// TIA Portal project "Sistema_de_silos" (V16) (continued)
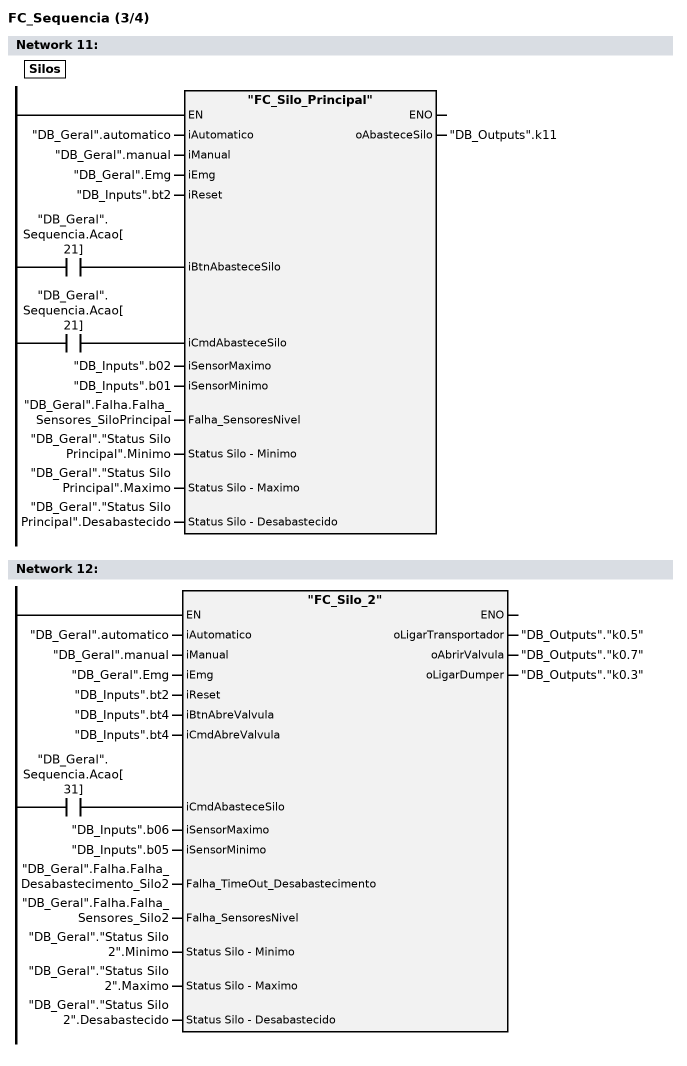
   Label( Silos )
   RUNG wire#powerrail
      "FC_Silo_Principal"(iBtnAbasteceSilo := wire#w1, iCmdAbasteceSilo := wire#w2, iAutomatico := "DB_Geral".automatico, iManual := "DB_Geral".manual, iEmg := "DB_Geral".Emg, iReset := "DB_Inputs".bt2, iSensorMaximo := "DB_Inputs".b02, iSensorMinimo := "DB_Inputs".b01, Falha_SensoresNivel := "DB_Geral".Falha.Falha_Sensores_SiloPrincipal, "Status Silo - Minimo" := "DB_Geral"."Status Silo Principal".Minimo, "Status Silo - Maximo" := "DB_Geral"."Status Silo Principal".Maximo, "Status Silo - Desabastecido" := "DB_Geral"."Status Silo Principal".Desabastecido, oAbasteceSilo => "DB_Outputs".k11)
   END_RUNG
   RUNG wire#powerrail
      Contact( "DB_Geral".Sequencia.Acao[21] )
   END_RUNG wire#w1
   RUNG wire#powerrail
      Contact( "DB_Geral".Sequencia.Acao[21] )
   END_RUNG wire#w2
   // the same network as SCL:
   Silos:
   "FC_Silo_Principal"(iAutomatico := "DB_Geral".automatico,
                       iManual := "DB_Geral".manual,
                       iEmg := "DB_Geral".Emg,
                       iReset := "DB_Inputs".bt2,
                       iBtnAbasteceSilo := "DB_Geral".Sequencia.Acao[21],
                       iCmdAbasteceSilo := "DB_Geral".Sequencia.Acao[21],
                       iSensorMaximo := "DB_Inputs".b02,
                       iSensorMinimo := "DB_Inputs".b01,
                       Falha_SensoresNivel := "DB_Geral".Falha.Falha_Sensores_SiloPrincipal,
                       "Status Silo - Minimo" := "DB_Geral"."Status Silo Principal".Minimo,
                       "Status Silo - Maximo" := "DB_Geral"."Status Silo Principal".Maximo,
                       "Status Silo - Desabastecido" := "DB_Geral"."Status Silo Principal".Desabastecido,
                       oAbasteceSilo => "DB_Outputs".k11);
END_REGION

REGION Network 12
   RUNG wire#powerrail
      "FC_Silo_2"(iCmdAbasteceSilo := wire#w1, iAutomatico := "DB_Geral".automatico, iManual := "DB_Geral".manual, iEmg := "DB_Geral".Emg, iReset := "DB_Inputs".bt2, iBtnAbreValvula := "DB_Inputs".bt4, iCmdAbreValvula := "DB_Inputs".bt4, iSensorMaximo := "DB_Inputs".b06, iSensorMinimo := "DB_Inputs".b05, Falha_TimeOut_Desabastecimento := "DB_Geral".Falha.Falha_Desabastecimento_Silo2, Falha_SensoresNivel := "DB_Geral".Falha.Falha_Sensores_Silo2, "Status Silo - Minimo" := "DB_Geral"."Status Silo 2".Minimo, "Status Silo - Maximo" := "DB_Geral"."Status Silo 2".Maximo, "Status Silo - Desabastecido" := "DB_Geral"."Status Silo 2".Desabastecido, oLigarTransportador => "DB_Outputs"."k0.5", oAbrirValvula => "DB_Outputs"."k0.7", oLigarDumper => "DB_Outputs"."k0.3")
   END_RUNG
   RUNG wire#powerrail
      Contact( "DB_Geral".Sequencia.Acao[31] )
   END_RUNG wire#w1
   // the same network as SCL:
   "FC_Silo_2"(iAutomatico := "DB_Geral".automatico,
               iManual := "DB_Geral".manual,
               iEmg := "DB_Geral".Emg,
               iReset := "DB_Inputs".bt2,
               iBtnAbreValvula := "DB_Inputs".bt4,
               iCmdAbreValvula := "DB_Inputs".bt4,
               iCmdAbasteceSilo := "DB_Geral".Sequencia.Acao[31],
               iSensorMaximo := "DB_Inputs".b06,
               iSensorMinimo := "DB_Inputs".b05,
               Falha_TimeOut_Desabastecimento := "DB_Geral".Falha.Falha_Desabastecimento_Silo2,
               Falha_SensoresNivel := "DB_Geral".Falha.Falha_Sensores_Silo2,
               "Status Silo - Minimo" := "DB_Geral"."Status Silo 2".Minimo,
               "Status Silo - Maximo" := "DB_Geral"."Status Silo 2".Maximo,
               "Status Silo - Desabastecido" := "DB_Geral"."Status Silo 2".Desabastecido,
               oLigarTransportador => "DB_Outputs"."k0.5",
               oAbrirValvula => "DB_Outputs"."k0.7",
               oLigarDumper => "DB_Outputs"."k0.3");
END_REGION

REGION Network 13
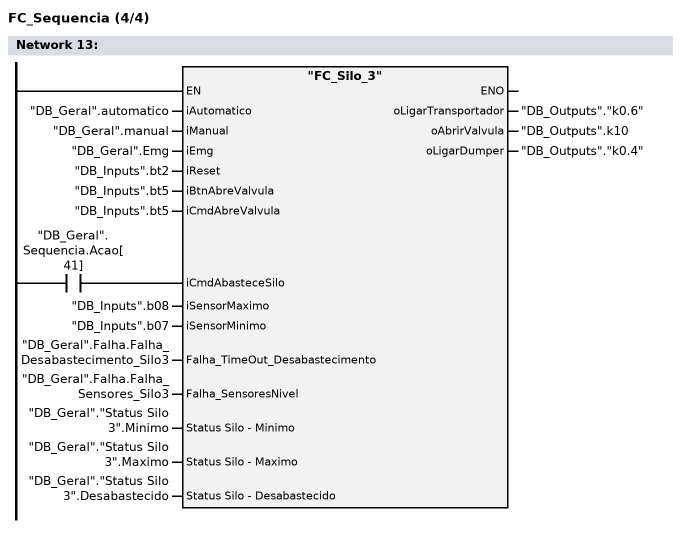
   RUNG wire#powerrail
      "FC_Silo_3"(iCmdAbasteceSilo := wire#w1, iAutomatico := "DB_Geral".automatico, iManual := "DB_Geral".manual, iEmg := "DB_Geral".Emg, iReset := "DB_Inputs".bt2, iBtnAbreValvula := "DB_Inputs".bt5, iCmdAbreValvula := "DB_Inputs".bt5, iSensorMaximo := "DB_Inputs".b08, iSensorMinimo := "DB_Inputs".b07, Falha_TimeOut_Desabastecimento := "DB_Geral".Falha.Falha_Desabastecimento_Silo3, Falha_SensoresNivel := "DB_Geral".Falha.Falha_Sensores_Silo3, "Status Silo - Minimo" := "DB_Geral"."Status Silo 3".Minimo, "Status Silo - Maximo" := "DB_Geral"."Status Silo 3".Maximo, "Status Silo - Desabastecido" := "DB_Geral"."Status Silo 3".Desabastecido, oLigarTransportador => "DB_Outputs"."k0.6", oAbrirValvula => "DB_Outputs".k10, oLigarDumper => "DB_Outputs"."k0.4")
   END_RUNG
   RUNG wire#powerrail
      Contact( "DB_Geral".Sequencia.Acao[41] )
   END_RUNG wire#w1
   // the same network as SCL:
   "FC_Silo_3"(iAutomatico := "DB_Geral".automatico,
               iManual := "DB_Geral".manual,
               iEmg := "DB_Geral".Emg,
               iReset := "DB_Inputs".bt2,
               iBtnAbreValvula := "DB_Inputs".bt5,
               iCmdAbreValvula := "DB_Inputs".bt5,
               iCmdAbasteceSilo := "DB_Geral".Sequencia.Acao[41],
               iSensorMaximo := "DB_Inputs".b08,
               iSensorMinimo := "DB_Inputs".b07,
               Falha_TimeOut_Desabastecimento := "DB_Geral".Falha.Falha_Desabastecimento_Silo3,
               Falha_SensoresNivel := "DB_Geral".Falha.Falha_Sensores_Silo3,
               "Status Silo - Minimo" := "DB_Geral"."Status Silo 3".Minimo,
               "Status Silo - Maximo" := "DB_Geral"."Status Silo 3".Maximo,
               "Status Silo - Desabastecido" := "DB_Geral"."Status Silo 3".Desabastecido,
               oLigarTransportador => "DB_Outputs"."k0.6",
               oAbrirValvula => "DB_Outputs".k10,
               oLigarDumper => "DB_Outputs"."k0.4");
END_REGION
END_FUNCTION

FUNCTION "FC_Silo_2" : Void   // FC5, LAD
{ S7_Optimized_Access := 'TRUE' }
VERSION : 0.1
   VAR_INPUT
      iAutomatico : Bool;
      iManual : Bool;
      iEmg : Bool;
      iReset : Bool;
      iBtnAbreValvula : Bool;
      iCmdAbreValvula : Bool;
      iCmdAbasteceSilo : Bool;
      iSensorMaximo : Bool;
      iSensorMinimo : Bool;
   END_VAR
   VAR_OUTPUT
      oLigarTransportador : Bool;
      oAbrirValvula : Bool;
      oLigarDumper : Bool;
   END_VAR
   VAR_IN_OUT
      Falha_TimeOut_Desabastecimento : Bool;
      Falha_SensoresNivel : Bool;
      "Status Silo - Minimo" : Bool;
      "Status Silo - Maximo" : Bool;
      "Status Silo - Desabastecido" : Bool;
   END_VAR
   VAR CONSTANT
      Velocidade_fluxo : Int := 12;
   END_VAR
BEGIN

REGION Network 1
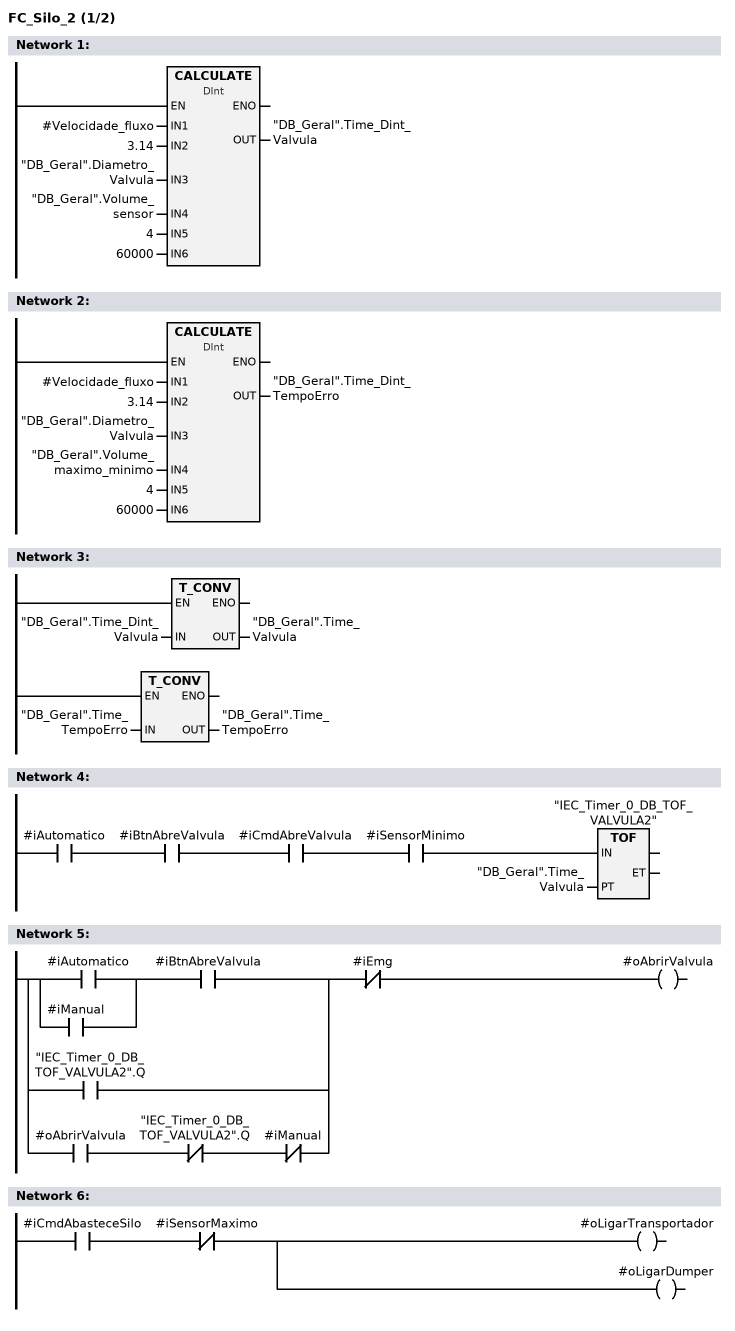
   RUNG wire#powerrail
      { S7_Templates := "SrcType := DInt"; S7_Expression := "(IN4 / (IN1* ((IN2*IN3*IN3) / IN5))) * IN6" } Calculate(in1 := #Velocidade_fluxo, in2 := 3.14, in3 := "DB_Geral".Diametro_Valvula, in4 := "DB_Geral".Volume_sensor, in5 := 4, in6 := 60000, out => "DB_Geral".Time_Dint_Valvula)
   END_RUNG
   // the same network as SCL:
   "DB_Geral".Time_Dint_Valvula := ("DB_Geral".Volume_sensor / (#Velocidade_fluxo* ((3.14*"DB_Geral".Diametro_Valvula*"DB_Geral".Diametro_Valvula) / 4))) * 60000;
END_REGION

REGION Network 2
   RUNG wire#powerrail
      { S7_Templates := "SrcType := DInt"; S7_Expression := "(IN4 / (IN1* ((IN2*IN3*IN3) / IN5))) * IN6" } Calculate(in1 := #Velocidade_fluxo, in2 := 3.14, in3 := "DB_Geral".Diametro_Valvula, in4 := "DB_Geral".Volume_maximo_minimo, in5 := 4, in6 := 60000, out => "DB_Geral".Time_Dint_TempoErro)
   END_RUNG
   // the same network as SCL:
   "DB_Geral".Time_Dint_TempoErro := ("DB_Geral".Volume_maximo_minimo / (#Velocidade_fluxo* ((3.14*"DB_Geral".Diametro_Valvula*"DB_Geral".Diametro_Valvula) / 4))) * 60000;
END_REGION

REGION Network 3
   "DB_Geral".Time_Valvula := T_CONV(IN := "DB_Geral".Time_Dint_Valvula);
   "DB_Geral".Time_TempoErro := T_CONV(IN := "DB_Geral".Time_TempoErro);
END_REGION

REGION Network 4
   "IEC_Timer_0_DB_TOF_VALVULA2".TOF(IN := #iAutomatico AND #iBtnAbreValvula AND #iCmdAbreValvula AND #iSensorMinimo,
                           PT := "DB_Geral".Time_Valvula);
END_REGION

REGION Network 5
   RUNG wire#powerrail
      Contact( #iAutomatico )
      wire#w1
      Contact( #iBtnAbreValvula )
      wire#w2
      I_Contact( #iEmg )
      Coil( #oAbrirValvula )
   END_RUNG
   RUNG wire#powerrail
      Contact( #iManual )
   END_RUNG wire#w1
   RUNG wire#powerrail
      Contact( "IEC_Timer_0_DB_TOF_VALVULA2".Q )
   END_RUNG wire#w2
   RUNG wire#powerrail
      Contact( #oAbrirValvula )
      I_Contact( "IEC_Timer_0_DB_TOF_VALVULA2".Q )
      I_Contact( #iManual )
   END_RUNG wire#w2
   // the same network as SCL:
   #oAbrirValvula := (((#iAutomatico OR #iManual) AND #iBtnAbreValvula) OR "IEC_Timer_0_DB_TOF_VALVULA2".Q OR (#oAbrirValvula AND NOT "IEC_Timer_0_DB_TOF_VALVULA2".Q AND NOT #iManual)) AND NOT #iEmg;
END_REGION

REGION Network 6
   RUNG wire#powerrail
      Contact( #iCmdAbasteceSilo )
      I_Contact( #iSensorMaximo )
      wire#w1
      Coil( #oLigarTransportador )
   END_RUNG
   RUNG wire#w1
      Coil( #oLigarDumper )
   END_RUNG
   // the same network as SCL:
   #oLigarTransportador := #iCmdAbasteceSilo AND NOT #iSensorMaximo;
   #oLigarDumper := #oLigarTransportador;
END_REGION

REGION Network 7: Silo Principal - Reserva do produto
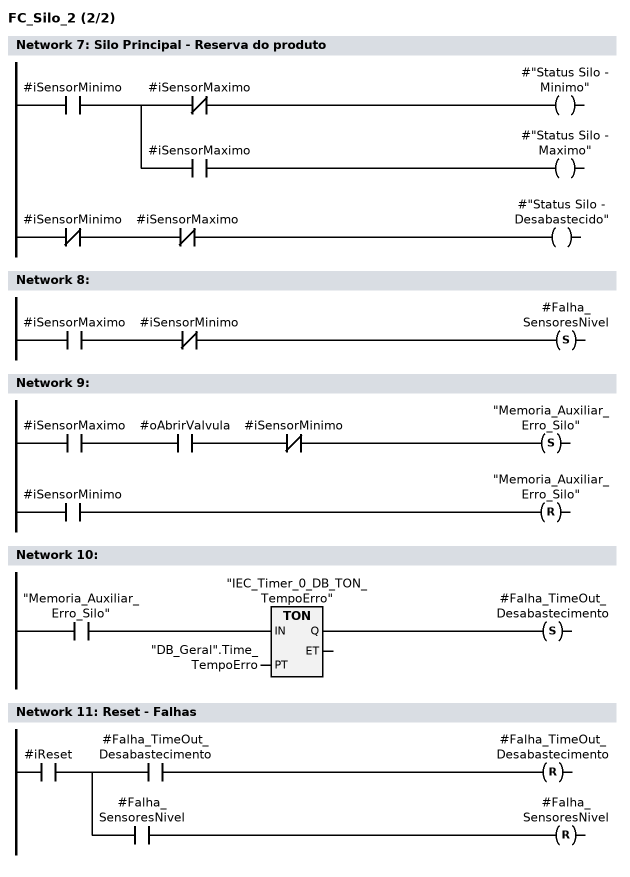
   RUNG wire#powerrail
      Contact( #iSensorMinimo )
      wire#w1
      I_Contact( #iSensorMaximo )
      Coil( #"Status Silo - Minimo" )
   END_RUNG
   RUNG wire#w1
      Contact( #iSensorMaximo )
      Coil( #"Status Silo - Maximo" )
   END_RUNG
   RUNG wire#powerrail
      I_Contact( #iSensorMinimo )
      I_Contact( #iSensorMaximo )
      Coil( #"Status Silo - Desabastecido" )
   END_RUNG
   // the same network as SCL:
   #"Status Silo - Minimo" := #iSensorMinimo AND NOT #iSensorMaximo;
   #"Status Silo - Maximo" := #iSensorMinimo AND #iSensorMaximo;
   #"Status Silo - Desabastecido" := NOT #iSensorMinimo AND NOT #iSensorMaximo;
END_REGION

REGION Network 8
   RUNG wire#powerrail
      Contact( #iSensorMaximo )
      I_Contact( #iSensorMinimo )
      S_Coil( #Falha_SensoresNivel )
   END_RUNG
   // the same network as SCL:
   IF #iSensorMaximo AND NOT #iSensorMinimo THEN #Falha_SensoresNivel := TRUE; END_IF;
END_REGION

REGION Network 9
   RUNG wire#powerrail
      Contact( #iSensorMaximo )
      Contact( #oAbrirValvula )
      I_Contact( #iSensorMinimo )
      S_Coil( "Memoria_Auxiliar_Erro_Silo" )
   END_RUNG
   RUNG wire#powerrail
      Contact( #iSensorMinimo )
      R_Coil( "Memoria_Auxiliar_Erro_Silo" )
   END_RUNG
   // the same network as SCL:
   IF #iSensorMaximo AND #oAbrirValvula AND NOT #iSensorMinimo THEN
       "Memoria_Auxiliar_Erro_Silo" := TRUE;
   END_IF;
   IF #iSensorMinimo THEN "Memoria_Auxiliar_Erro_Silo" := FALSE; END_IF;
END_REGION

REGION Network 10
   "IEC_Timer_0_DB_TON_TempoErro".TON(IN := "Memoria_Auxiliar_Erro_Silo", PT := "DB_Geral".Time_TempoErro);
   IF "IEC_Timer_0_DB_TON_TempoErro".Q THEN #Falha_TimeOut_Desabastecimento := TRUE; END_IF;
END_REGION

REGION Network 11: Reset - Falhas
   RUNG wire#powerrail
      Contact( #iReset )
      wire#w1
      Contact( #Falha_TimeOut_Desabastecimento )
      R_Coil( #Falha_TimeOut_Desabastecimento )
   END_RUNG
   RUNG wire#w1
      Contact( #Falha_SensoresNivel )
      R_Coil( #Falha_SensoresNivel )
   END_RUNG
   // the same network as SCL:
   IF #iReset AND #Falha_TimeOut_Desabastecimento THEN #Falha_TimeOut_Desabastecimento := FALSE; END_IF;
   IF #iReset AND #Falha_SensoresNivel THEN #Falha_SensoresNivel := FALSE; END_IF;
END_REGION
END_FUNCTION

FUNCTION "FC_Silo_Principal" : Void   // FC6, LAD
{ S7_Optimized_Access := 'TRUE' }
VERSION : 0.1
   VAR_INPUT
      iAutomatico : Bool;
      iManual : Bool;
      iEmg : Bool;
      iReset : Bool;
      iBtnAbasteceSilo : Bool;
      iCmdAbasteceSilo : Bool;
      iSensorMaximo : Bool;
      iSensorMinimo : Bool;
   END_VAR
   VAR_OUTPUT
      oAbasteceSilo : Bool;
   END_VAR
   VAR_IN_OUT
      Falha_SensoresNivel : Bool;
      "Status Silo - Minimo" : Bool;
      "Status Silo - Maximo" : Bool;
      "Status Silo - Desabastecido" : Bool;
   END_VAR
BEGIN

REGION Network 1
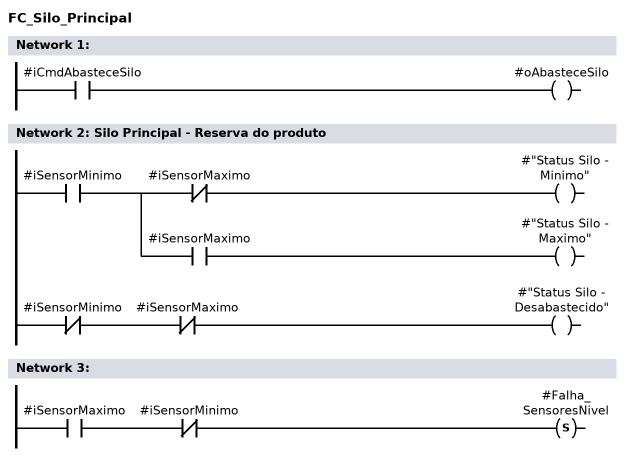
   RUNG wire#powerrail
      Contact( #iCmdAbasteceSilo )
      Coil( #oAbasteceSilo )
   END_RUNG
   // the same network as SCL:
   #oAbasteceSilo := #iCmdAbasteceSilo;
END_REGION

REGION Network 2: Silo Principal - Reserva do produto
   RUNG wire#powerrail
      Contact( #iSensorMinimo )
      wire#w1
      I_Contact( #iSensorMaximo )
      Coil( #"Status Silo - Minimo" )
   END_RUNG
   RUNG wire#w1
      Contact( #iSensorMaximo )
      Coil( #"Status Silo - Maximo" )
   END_RUNG
   RUNG wire#powerrail
      I_Contact( #iSensorMinimo )
      I_Contact( #iSensorMaximo )
      Coil( #"Status Silo - Desabastecido" )
   END_RUNG
   // the same network as SCL:
   #"Status Silo - Minimo" := #iSensorMinimo AND NOT #iSensorMaximo;
   #"Status Silo - Maximo" := #iSensorMinimo AND #iSensorMaximo;
   #"Status Silo - Desabastecido" := NOT #iSensorMinimo AND NOT #iSensorMaximo;
END_REGION

REGION Network 3
   RUNG wire#powerrail
      Contact( #iSensorMaximo )
      I_Contact( #iSensorMinimo )
      S_Coil( #Falha_SensoresNivel )
   END_RUNG
   // the same network as SCL:
   IF #iSensorMaximo AND NOT #iSensorMinimo THEN #Falha_SensoresNivel := TRUE; END_IF;
END_REGION
END_FUNCTION

FUNCTION "FC_Silo_3" : Void   // FC7, LAD
{ S7_Optimized_Access := 'TRUE' }
VERSION : 0.1
   VAR_INPUT
      iAutomatico : Bool;
      iManual : Bool;
      iEmg : Bool;
      iReset : Bool;
      iBtnAbreValvula : Bool;
      iCmdAbreValvula : Bool;
      iCmdAbasteceSilo : Bool;
      iSensorMaximo : Bool;
      iSensorMinimo : Bool;
   END_VAR
   VAR_OUTPUT
      oLigarTransportador : Bool;
      oAbrirValvula : Bool;
      oLigarDumper : Bool;
   END_VAR
   VAR_IN_OUT
      Falha_TimeOut_Desabastecimento : Bool;
      Falha_SensoresNivel : Bool;
      "Status Silo - Minimo" : Bool;
      "Status Silo - Maximo" : Bool;
      "Status Silo - Desabastecido" : Bool;
   END_VAR
   VAR CONSTANT
      Velocidade_fluxo : Int := 12;
   END_VAR
BEGIN

REGION Network 1
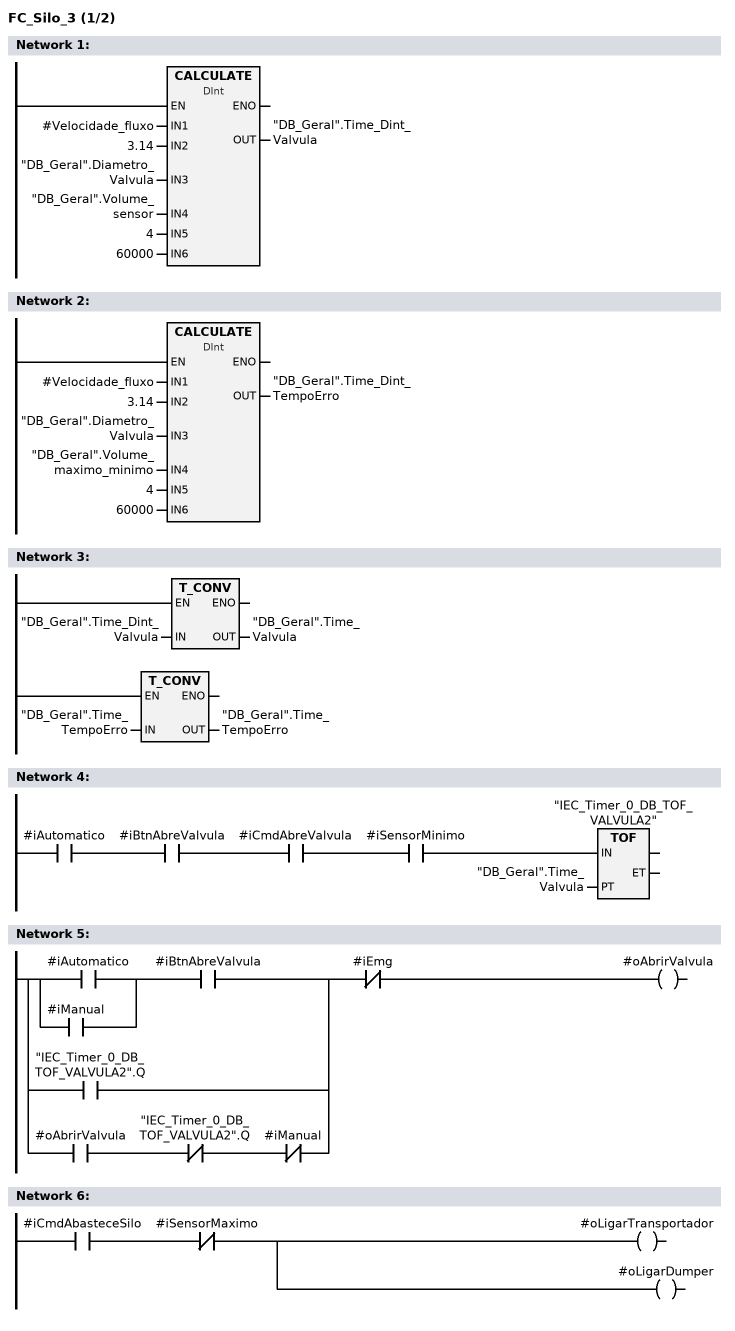
   RUNG wire#powerrail
      { S7_Templates := "SrcType := DInt"; S7_Expression := "(IN4 / (IN1* ((IN2*IN3*IN3) / IN5))) * IN6" } Calculate(in1 := #Velocidade_fluxo, in2 := 3.14, in3 := "DB_Geral".Diametro_Valvula, in4 := "DB_Geral".Volume_sensor, in5 := 4, in6 := 60000, out => "DB_Geral".Time_Dint_Valvula)
   END_RUNG
   // the same network as SCL:
   "DB_Geral".Time_Dint_Valvula := ("DB_Geral".Volume_sensor / (#Velocidade_fluxo* ((3.14*"DB_Geral".Diametro_Valvula*"DB_Geral".Diametro_Valvula) / 4))) * 60000;
END_REGION

REGION Network 2
   RUNG wire#powerrail
      { S7_Templates := "SrcType := DInt"; S7_Expression := "(IN4 / (IN1* ((IN2*IN3*IN3) / IN5))) * IN6" } Calculate(in1 := #Velocidade_fluxo, in2 := 3.14, in3 := "DB_Geral".Diametro_Valvula, in4 := "DB_Geral".Volume_maximo_minimo, in5 := 4, in6 := 60000, out => "DB_Geral".Time_Dint_TempoErro)
   END_RUNG
   // the same network as SCL:
   "DB_Geral".Time_Dint_TempoErro := ("DB_Geral".Volume_maximo_minimo / (#Velocidade_fluxo* ((3.14*"DB_Geral".Diametro_Valvula*"DB_Geral".Diametro_Valvula) / 4))) * 60000;
END_REGION

REGION Network 3
   "DB_Geral".Time_Valvula := T_CONV(IN := "DB_Geral".Time_Dint_Valvula);
   "DB_Geral".Time_TempoErro := T_CONV(IN := "DB_Geral".Time_TempoErro);
END_REGION

REGION Network 4
   "IEC_Timer_0_DB_TOF_VALVULA2".TOF(IN := #iAutomatico AND #iBtnAbreValvula AND #iCmdAbreValvula AND #iSensorMinimo,
                           PT := "DB_Geral".Time_Valvula);
END_REGION

REGION Network 5
   RUNG wire#powerrail
      Contact( #iAutomatico )
      wire#w1
      Contact( #iBtnAbreValvula )
      wire#w2
      I_Contact( #iEmg )
      Coil( #oAbrirValvula )
   END_RUNG
   RUNG wire#powerrail
      Contact( #iManual )
   END_RUNG wire#w1
   RUNG wire#powerrail
      Contact( "IEC_Timer_0_DB_TOF_VALVULA2".Q )
   END_RUNG wire#w2
   RUNG wire#powerrail
      Contact( #oAbrirValvula )
      I_Contact( "IEC_Timer_0_DB_TOF_VALVULA2".Q )
      I_Contact( #iManual )
   END_RUNG wire#w2
   // the same network as SCL:
   #oAbrirValvula := (((#iAutomatico OR #iManual) AND #iBtnAbreValvula) OR "IEC_Timer_0_DB_TOF_VALVULA2".Q OR (#oAbrirValvula AND NOT "IEC_Timer_0_DB_TOF_VALVULA2".Q AND NOT #iManual)) AND NOT #iEmg;
END_REGION

REGION Network 6
   RUNG wire#powerrail
      Contact( #iCmdAbasteceSilo )
      I_Contact( #iSensorMaximo )
      wire#w1
      Coil( #oLigarTransportador )
   END_RUNG
   RUNG wire#w1
      Coil( #oLigarDumper )
   END_RUNG
   // the same network as SCL:
   #oLigarTransportador := #iCmdAbasteceSilo AND NOT #iSensorMaximo;
   #oLigarDumper := #oLigarTransportador;
END_REGION

REGION Network 7: Silo Principal - Reserva do produto
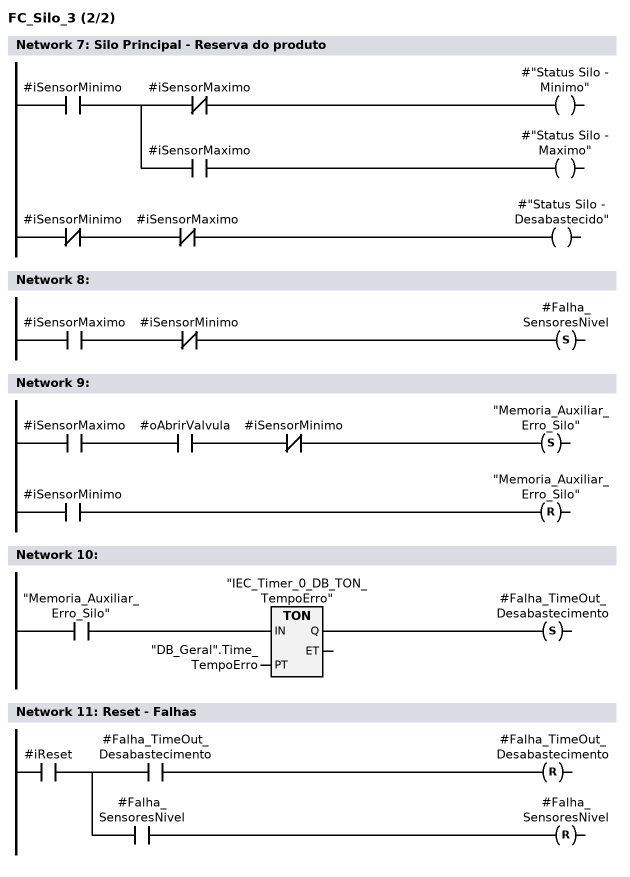
   RUNG wire#powerrail
      Contact( #iSensorMinimo )
      wire#w1
      I_Contact( #iSensorMaximo )
      Coil( #"Status Silo - Minimo" )
   END_RUNG
   RUNG wire#w1
      Contact( #iSensorMaximo )
      Coil( #"Status Silo - Maximo" )
   END_RUNG
   RUNG wire#powerrail
      I_Contact( #iSensorMinimo )
      I_Contact( #iSensorMaximo )
      Coil( #"Status Silo - Desabastecido" )
   END_RUNG
   // the same network as SCL:
   #"Status Silo - Minimo" := #iSensorMinimo AND NOT #iSensorMaximo;
   #"Status Silo - Maximo" := #iSensorMinimo AND #iSensorMaximo;
   #"Status Silo - Desabastecido" := NOT #iSensorMinimo AND NOT #iSensorMaximo;
END_REGION

REGION Network 8
   RUNG wire#powerrail
      Contact( #iSensorMaximo )
      I_Contact( #iSensorMinimo )
      S_Coil( #Falha_SensoresNivel )
   END_RUNG
   // the same network as SCL:
   IF #iSensorMaximo AND NOT #iSensorMinimo THEN #Falha_SensoresNivel := TRUE; END_IF;
END_REGION

REGION Network 9
   RUNG wire#powerrail
      Contact( #iSensorMaximo )
      Contact( #oAbrirValvula )
      I_Contact( #iSensorMinimo )
      S_Coil( "Memoria_Auxiliar_Erro_Silo" )
   END_RUNG
   RUNG wire#powerrail
      Contact( #iSensorMinimo )
      R_Coil( "Memoria_Auxiliar_Erro_Silo" )
   END_RUNG
   // the same network as SCL:
   IF #iSensorMaximo AND #oAbrirValvula AND NOT #iSensorMinimo THEN
       "Memoria_Auxiliar_Erro_Silo" := TRUE;
   END_IF;
   IF #iSensorMinimo THEN "Memoria_Auxiliar_Erro_Silo" := FALSE; END_IF;
END_REGION

REGION Network 10
   "IEC_Timer_0_DB_TON_TempoErro".TON(IN := "Memoria_Auxiliar_Erro_Silo", PT := "DB_Geral".Time_TempoErro);
   IF "IEC_Timer_0_DB_TON_TempoErro".Q THEN #Falha_TimeOut_Desabastecimento := TRUE; END_IF;
END_REGION

REGION Network 11: Reset - Falhas
   RUNG wire#powerrail
      Contact( #iReset )
      wire#w1
      Contact( #Falha_TimeOut_Desabastecimento )
      R_Coil( #Falha_TimeOut_Desabastecimento )
   END_RUNG
   RUNG wire#w1
      Contact( #Falha_SensoresNivel )
      R_Coil( #Falha_SensoresNivel )
   END_RUNG
   // the same network as SCL:
   IF #iReset AND #Falha_TimeOut_Desabastecimento THEN #Falha_TimeOut_Desabastecimento := FALSE; END_IF;
   IF #iReset AND #Falha_SensoresNivel THEN #Falha_SensoresNivel := FALSE; END_IF;
END_REGION
END_FUNCTION

ORGANIZATION_BLOCK "Main"   // OB1, LAD, ProgramCycle
TITLE = "Main Program Sweep (Cycle)"
{ S7_Optimized_Access := 'TRUE' }
VERSION : 0.1
   VAR_INPUT
      Initial_Call : Bool;   // Initial call of this OB
      Remanence : Bool;   // =True, if remanent data are available
   END_VAR
BEGIN
END_ORGANIZATION_BLOCK

(* ===== HMI "HMI_RT_1" =====
system functions are stored by id; their names below are inferred from use
connection "HMI_Connection_1": ETHERNET, S7_1200_OMS
connection "HMI_Connection_2": IF1 B, S7_1200_OMS
connection "HMI_Connection_3": IF1 B, S7_1200_OMS

HMI tags "Default tag table"
   "Tag_ScreenNumber" : UInt, internal

screen "Root screen" 1280x740, template "Template_1"
   on GenerateScreen: SetTag("Tag_ScreenNumber", 1)
   Button "HmiScreenItemData" at 79,35 size 213x73; TextOff 'Teste Screen'; PictureOff "Navigates to Teste Screen for TP1200 Comfort 16.0.0.0"; PictureOn "Navigates to Teste Screen for TP1200 Comfort 16.0.0.0"
      on Release: ActivateScreen("Teste Screen", 0)
   Button "HmiScreenItemData_1" at 1002,36 size 213x73; TextOff 'Operation Screen'; PictureOff "Navigates to Operation Screen for TP1200 Comfort 16.0.0.0"; PictureOn "Navigates to Operation Screen for TP1200 Comfort 16.0.0.0"
      on Release: ActivateScreen("Operation Screen", 0)
   Button "HmiScreenItemData_2" at 692,33 size 213x73; TextOff 'Fail/Emg Screen'; PictureOff "Navigates to Fail/Emg Screen for TP1200 Comfort 16.0.0.0"; PictureOn "Navigates to Fail/Emg Screen for TP1200 Comfort 16.0.0.0"
      on Release: ActivateScreen("Fail/Emg Screen", 0)
   Button "HmiScreenItemData_4" at 377,35 size 213x73; TextOff 'System screens'; PictureOff "Navigates to System screens for TP1200 Comfort 16.0.0.0"; PictureOn "Navigates to System screens for TP1200 Comfort 16.0.0.0"
      on Release: ActivateScreen("System screens", 0)
   GraphicView "Graphic view_3" at 361,257 size 541x174; Picture "Siemens Logo"

Template "Template_1" 1280x740
   Button "Exit" at 1200,679 size 78x59; TextOff 'Exit'; PictureOff "ExitRuntime_TP1200_Comfort_TR"; PictureOn "ExitRuntime_TP1200_Comfort_TR"
      on Release: StopRuntime(0)
   Button "Template_Button" at 1120,679 size 78x59; TextOff 'Text'
   Button "Template_Button_1" at 1040,679 size 78x59; TextOff 'Text'
   Button "Template_Button_2" at 960,679 size 78x59; TextOff 'Text'
   Button "Template_Button_3" at 880,679 size 78x59; TextOff 'Text'
   Button "Template_Button_4" at 800,679 size 78x59; TextOff 'Text'
   Button "Template_Button_5" at 720,679 size 78x59; TextOff 'Text'
   Button "Template_Button_6" at 640,679 size 78x59; TextOff 'Text'
   Button "Template_Button_7" at 561,679 size 78x59; TextOff 'Text'
   Button "Template_Button_8" at 481,679 size 78x59; TextOff 'Text'
   Button "Template_Button_9" at 401,679 size 78x59; TextOff 'Text'
   Button "Template_Button_10" at 321,679 size 78x59; TextOff 'Text'
   Button "Template_Button_11" at 241,679 size 78x59; TextOff 'Text'
   Button "Template_Button_12" at 161,679 size 78x59; TextOff 'Text'
   Button "Alarms" at 81,679 size 78x59; TextOff 'Alarms'; PictureOff "AlarmDisplay_TP1200_Comfort_TR"; PictureOn "AlarmDisplay_TP1200_Comfort_TR"
      on Release: function_ef3f5d25("Alarm window_Unacknowledged", -1)
   Button "Start screen" at 1,679 size 78x59; TextOff 'Start screen'; PictureOff "NavigateHome_TP1200_Comfort_TR"; PictureOn "NavigateHome_TP1200_Comfort_TR"
      on Release: ActivateScreen("Root screen", 0)

screen "Teste Screen" 1280x740, template "Template_1"
   on GenerateScreen: SetTag("Tag_ScreenNumber", 2)
   Button "Back" at 0,24 size 159x47; TextOff 'Back'
      on Release: ActivateScreen("Root screen", 0)
   Button "Button_1" at 10,127 size 200x95; TextOff 'Manual'
   Button "Button_2" at 9,271 size 200x95; TextOff 'Automatico'
   Button "Button_3" at 10,417 size 200x95; TextOff 'Emergência'
   Button "Button_4" at 11,563 size 200x95; TextOff 'Reset'
   Button "Button_5" at 1055,127 size 200x95; TextOff 'Valvula 1'
   Button "Button_6" at 1055,271 size 200x95; TextOff 'Valvula 2'

screen "Operation Screen" 1280x740, template "Template_1"
   on GenerateScreen: SetTag("Tag_ScreenNumber", 3)
   TextField "HmiScreenItemData" at 128,324 size 1024x27; Text 'Operation Screen'
   Button "Back" at 1,1 size 159x47; TextOff 'Back'
      on Release: ActivateScreen("Root screen", 0)

screen "Fail/Emg Screen" 1280x740, template "Template_1"
   on GenerateScreen: SetTag("Tag_ScreenNumber", 4)
   TextField "HmiScreenItemData" at 128,324 size 1024x27; Text 'Fail/Emg Screen'
   Button "Back" at 1,1 size 159x47; TextOff 'Back'
      on Release: ActivateScreen("Root screen", 0)

screen "System screens" 1280x740, template "Template_1"
   on GenerateScreen: SetTag("Tag_ScreenNumber", 5)
   Button "Back" at 1,1 size 159x47; TextOff 'Back'
      on Release: ActivateScreen("Root screen", 0)
   Button "HmiScreenItemData" at 36,95 size 159x47; TextOff 'SIMATIC PLC system diagnos...'; PictureOff "Navigates to SIMATIC PLC system diagnostics for TP1200 Comfort 16.0.0.0"; PictureOn "Navigates to SIMATIC PLC system diagnostics for TP1200 Comfort 16.0.0.0"
      on Release: ActivateScreen("SIMATIC PLC system diagnostics", 0)
   Button "HmiScreenItemData_1" at 36,154 size 159x47; TextOff 'System settings'; PictureOff "Navigates to System settings for TP1200 Comfort 16.0.0.0"; PictureOn "Navigates to System settings for TP1200 Comfort 16.0.0.0"
      on Release: ActivateScreen("System settings", 0)
   Button "HmiScreenItemData_2" at 36,213 size 159x47; TextOff 'System information'; PictureOff "Navigates to System information for TP1200 Comfort 16.0.0.0"; PictureOn "Navigates to System information for TP1200 Comfort 16.0.0.0"
      on Release: ActivateScreen("System information", 0)

screen "SIMATIC PLC system diagnostics" 1280x740, template "Template_1"
   on GenerateScreen: SetTag("Tag_ScreenNumber", 6)
   SysDiagControl "HmiScreenItemData" at 1,49 size 1276x623
   Button "Back" at 1,1 size 159x47; TextOff 'Back'
      on Release: ActivateScreen("System screens", 0)

screen "System settings" 1280x740, template "Template_1"
   on GenerateScreen: SetTag("Tag_ScreenNumber", 7)
   Button "Calibrate screen" at 36,95 size 159x47; TextOff 'Calibrate screen'
      on Release: function_bc3e350c()
   Button "Clean screen" at 36,154 size 159x47; TextOff 'Clean screen'
      on Release: function_be740847(30)
   Button "Back" at 1,1 size 159x47; TextOff 'Back'
      on Release: ActivateScreen("System screens", 0)

screen "System information" 1280x740, template "Template_1"
   on GenerateScreen: SetTag("Tag_ScreenNumber", 8)
   TextField "HmiScreenItemData" at 35,51 size 171x28; Text 'HMI device type:'
   TextField "HmiScreenItemData_1" at 241,51 size 1004x28; Text 'TP1200 Comfort 16.0.0.0'
   TextField "HmiScreenItemData_2" at 35,81 size 171x28; Text 'Version:'
   TextField "HmiScreenItemData_3" at 35,111 size 171x28; Text 'Connection:'
   TextField "HmiScreenItemData_4" at 241,111 size 1004x28; Text 'ETHERNET'
   TextField "HmiScreenItemData_5" at 35,141 size 171x28; Text 'PLC:'
   TextField "HmiScreenItemData_6" at 241,141 size 1004x28; Text 'SIMATIC S7 1200'
   Button "Display version" at 241,81 size 1004x28; TextOff 'Display version'
      on Release: function_febcb963(-1)
   Button "Back" at 1,1 size 159x47; TextOff 'Back'
      on Release: ActivateScreen("System screens", 0)
*)